
screen "0999_Service" 1280x800, template "Navigation"
   on GenerateScreen: SetTag("NavScreenChange", 5)
   on ClearScreen: SetTag("NavScreenChange", 0)
   Button "Button_3" at 326,104 size 451x32; TextOff 'Service'
   GraphicView "Graphic view_1" at 613,200 size 64x100; Picture "tank"
   GraphicView "Graphic view_2" at 385,180 size 144x140; Picture "Mcn"
   GraphicView "Graphic view_3" at 192,180 size 144x140; Picture "Machine"
   GraphicView "Graphic view_4" at 952,180 size 144x140; Picture "images_4"
   GraphicView "Graphic view_5" at 216,387 size 96x98; Picture "switch_off"
   GraphicView "Graphic view_6" at 781,224 size 116x60; Picture "Graphic_1"
   GraphicView "Graphic view_7" at 399,647 size 116x100; Picture "LARGESCALLEDVALUE"
   GraphicView "Graphic view_8" at 587,647 size 116x100; Picture "osiloskope_1"
   GraphicView "Graphic view_9" at 206,647 size 116x100; Picture "ethernet"
      Visibility <- "NavUserChange"
   Button "MixingHeadButton_1" at 565,182 size 160x136; TextOff 'Tank'; PictureOff "tank"
      on Click: ActivateScreen("0006_Tank", 0)
   Button "MixingHeadButton_3" at 944,182 size 160x136; TextOff 'Metering Pump'
      on Click: ActivateScreen("0004_Mixinghead", 0)
   Button "MixingHeadButton_2" at 184,182 size 160x136; TextOff 'General Machine'
      on Click: ActivateScreen("0021_Machine", 0)
   Button "MixingHeadButton_4" at 944,627 size 160x136; TextOff 'KM'; Authorization "User administration"
      Visibility <- "NavUserChange"
      on Click: ActivateScreen("2000_Configuration", 0)
   Button "MixingHeadButton_5" at 759,182 size 160x136; TextOff 'Mixinghead'
      on Click: ActivateScreen("0010_Pump", 0)
   Button "MixingHeadButton" at 377,182 size 160x136; TextOff 'Mixing Hydraulic'
      on Click: ActivateScreen("0002_MixingHeadHydraulic", 0)
   Button "MixingHeadButton_7" at 184,629 size 160x136; TextOff 'Network Setting'; Authorization "User administration"
      on Click: ActivateScreen("0014_Network Setting", 0)
      Visibility <- "NavUserChange"
   Button "MixingHeadButton_8" at 377,629 size 160x136; TextOff 'Large Scalled Values'
      on Click: ActivateScreen("0100_LargeScalledValues", 0); SetTag("NavScreenChange", 3); SetTag("LargeScalleValues Control", 1)
   Button "MixingHeadButton_9" at 565,629 size 160x136; TextOff 'Oscilloscope'
      on Click: ActivateScreen("0015_Oscilloscope", 0); SetTag("NavScreenChange", 2)
   Button "MixingHeadButton_10" at 184,368 size 160x136; TextOff 'Switch Menue'
      on Click: ActivateScreen("0009_Switch Menu", 0)
   Button "MixingHeadButton_11" at 759,623 size 160x136; TextOff 'Service & Solutions'
      on Click: ActivateScreen("9020_Service", 0)

screen "0016_Osciloscope Setting" 1280x800, template "Navigation"
   SymbolicIOField "Symbolic I/O field_11" at 704,218 size 160x30; TextOn '1'; TextOff '0'; TextList "oscilloscope_sensor_by_pump"
      Visibility <- "DB025_Oszilloskop_Graph{1}_Auswahl"
      ProcessValue <- "DB025_Oszilloskop_Graph{1}_Sensor"
   SymbolicIOField "Symbolic I/O field_15" at 704,270 size 160x30; TextOn '1'; TextOff '0'; TextList "oscilloscope_sensor_by_pump"
      Visibility <- "DB025_Oszilloskop_Graph{2}_Auswahl"
      ProcessValue <- "DB025_Oszilloskop_Graph{2}_Sensor"
   SymbolicIOField "Symbolic I/O field_19" at 704,322 size 160x30; TextOn '1'; TextOff '0'; TextList "oscilloscope_sensor_by_pump"
      ProcessValue <- "DB025_Oszilloskop_Graph{3}_Sensor"
      Visibility <- "DB025_Oszilloskop_Graph{3}_Auswahl"
   SymbolicIOField "Symbolic I/O field_23" at 704,374 size 160x30; TextOn '1'; TextOff '0'; TextList "oscilloscope_sensor_by_pump"
      ProcessValue <- "DB025_Oszilloskop_Graph{4}_Sensor"
      Visibility <- "DB025_Oszilloskop_Graph{4}_Auswahl"
   SymbolicIOField "Symbolic I/O field_27" at 704,426 size 160x30; TextOn '1'; TextOff '0'; TextList "oscilloscope_sensor_by_pump"
      ProcessValue <- "DB025_Oszilloskop_Graph{5}_Sensor"
      Visibility <- "DB025_Oszilloskop_Graph{5}_Auswahl"
   SymbolicIOField "Symbolic I/O field_31" at 704,478 size 160x30; TextOn '1'; TextOff '0'; TextList "oscilloscope_sensor_by_pump"
      ProcessValue <- "DB025_Oszilloskop_Graph{6}_Sensor"
      Visibility <- "DB025_Oszilloskop_Graph{6}_Auswahl"
   SymbolicIOField "Symbolic I/O field_35" at 704,530 size 160x30; TextOn '1'; TextOff '0'; TextList "oscilloscope_sensor_by_pump"
      ProcessValue <- "DB025_Oszilloskop_Graph{7}_Sensor"
      Visibility <- "DB025_Oszilloskop_Graph{7}_Auswahl"
   SymbolicIOField "Symbolic I/O field_39" at 704,582 size 160x30; TextOn '1'; TextOff '0'; TextList "oscilloscope_sensor_by_pump"
      ProcessValue <- "DB025_Oszilloskop_Graph{8}_Sensor"
      Visibility <- "DB025_Oszilloskop_Graph{8}_Auswahl"
   SymbolicIOField "Symbolic I/O field_12" at 704,218 size 160x30; TextOn '1'; TextOff '0'; TextList "oscilloscope_sensor_by_Tank"
      Visibility <- "DB025_Oszilloskop_Graph{1}_Auswahl"
      ProcessValue <- "DB025_Oszilloskop_Graph{1}_Sensor"
   SymbolicIOField "Symbolic I/O field_16" at 704,270 size 160x30; TextOn '1'; TextOff '0'; TextList "oscilloscope_sensor_by_Tank"
      Visibility <- "DB025_Oszilloskop_Graph{2}_Auswahl"
      ProcessValue <- "DB025_Oszilloskop_Graph{2}_Sensor"
   SymbolicIOField "Symbolic I/O field_20" at 704,322 size 160x30; TextOn '1'; TextOff '0'; TextList "oscilloscope_sensor_by_Tank"
      Visibility <- "DB025_Oszilloskop_Graph{3}_Auswahl"
      ProcessValue <- "DB025_Oszilloskop_Graph{3}_Sensor"
   SymbolicIOField "Symbolic I/O field_24" at 704,374 size 160x30; TextOn '1'; TextOff '0'; TextList "oscilloscope_sensor_by_Tank"
      Visibility <- "DB025_Oszilloskop_Graph{4}_Auswahl"
      ProcessValue <- "DB025_Oszilloskop_Graph{4}_Sensor"
   SymbolicIOField "Symbolic I/O field_28" at 704,426 size 160x30; TextOn '1'; TextOff '0'; TextList "oscilloscope_sensor_by_Tank"
      Visibility <- "DB025_Oszilloskop_Graph{5}_Auswahl"
      ProcessValue <- "DB025_Oszilloskop_Graph{5}_Sensor"
   SymbolicIOField "Symbolic I/O field_32" at 704,478 size 160x30; TextOn '1'; TextOff '0'; TextList "oscilloscope_sensor_by_Tank"
      Visibility <- "DB025_Oszilloskop_Graph{6}_Auswahl"
      ProcessValue <- "DB025_Oszilloskop_Graph{6}_Sensor"
   SymbolicIOField "Symbolic I/O field_36" at 704,530 size 160x30; TextOn '1'; TextOff '0'; TextList "oscilloscope_sensor_by_Tank"
      Visibility <- "DB025_Oszilloskop_Graph{7}_Auswahl"
      ProcessValue <- "DB025_Oszilloskop_Graph{7}_Sensor"
   SymbolicIOField "Symbolic I/O field_40" at 704,582 size 160x30; TextOn '1'; TextOff '0'; TextList "oscilloscope_sensor_by_Tank"
      Visibility <- "DB025_Oszilloskop_Graph{8}_Auswahl"
      ProcessValue <- "DB025_Oszilloskop_Graph{8}_Sensor"
   Button "Button_10" at 120,157 size 967x494; TextOff 'Text'
   Button "Button_3" at 326,104 size 451x32; TextOff 'Oscilloscope Settings'
   Button "Button_6" at 182,218 size 50x30; TextOff '1.'
   TextField "Text field_1" at 238,194 size 84x22; Text 'Selection'
   SymbolicIOField "Symbolic I/O field_1" at 238,218 size 160x30; TextOff '0'; TextOn '1'; TextList "oscilloscope_selection"
      ProcessValue <- "DB025_Oszilloskop_Graph{1}_Auswahl"
   Button "Button_1" at 182,270 size 50x30; TextOff '2.'
   TextField "Text field_2" at 238,246 size 84x22; Text 'Selection'
   SymbolicIOField "Symbolic I/O field_2" at 238,270 size 160x30; TextOn '1'; TextOff '0'; TextList "oscilloscope_selection"
      ProcessValue <- "DB025_Oszilloskop_Graph{2}_Auswahl"
   Button "Button_2" at 182,322 size 50x30; TextOff '3.'
   TextField "Text field_3" at 238,298 size 84x22; Text 'Selection'
   SymbolicIOField "Symbolic I/O field_3" at 238,322 size 160x30; TextOn '1'; TextOff '0'; TextList "oscilloscope_selection"
      ProcessValue <- "DB025_Oszilloskop_Graph{3}_Auswahl"
   Button "Button_4" at 182,374 size 50x30; TextOff '4.'
   TextField "Text field_4" at 238,350 size 84x22; Text 'Selection'
   SymbolicIOField "Symbolic I/O field_4" at 238,374 size 160x30; TextOn '1'; TextOff '0'; TextList "oscilloscope_selection"
      ProcessValue <- "DB025_Oszilloskop_Graph{4}_Auswahl"
   Button "Button_5" at 182,426 size 50x30; TextOff '5.'
   TextField "Text field_5" at 238,402 size 84x22; Text 'Selection'
   SymbolicIOField "Symbolic I/O field_5" at 238,426 size 160x30; TextOn '1'; TextOff '0'; TextList "oscilloscope_selection"
      ProcessValue <- "DB025_Oszilloskop_Graph{5}_Auswahl"
   Button "Button_7" at 182,478 size 50x30; TextOff '6.'
   TextField "Text field_6" at 238,454 size 84x22; Text 'Selection'
   SymbolicIOField "Symbolic I/O field_6" at 238,478 size 160x30; TextOn '1'; TextOff '0'; TextList "oscilloscope_selection"
      ProcessValue <- "DB025_Oszilloskop_Graph{6}_Auswahl"
   Button "Button_8" at 182,530 size 50x30; TextOff '7.'
   TextField "Text field_7" at 238,506 size 84x22; Text 'Selection'
   SymbolicIOField "Symbolic I/O field_7" at 238,530 size 160x30; TextOn '1'; TextOff '0'; TextList "oscilloscope_selection"
      ProcessValue <- "DB025_Oszilloskop_Graph{7}_Auswahl"
   Button "Button_9" at 182,582 size 50x30; TextOff '8.'
   TextField "Text field_8" at 238,558 size 84x22; Text 'Selection'
   SymbolicIOField "Symbolic I/O field_8" at 238,582 size 160x30; TextOn '1'; TextOff '0'; TextList "oscilloscope_selection"
      ProcessValue <- "DB025_Oszilloskop_Graph{8}_Auswahl"
   TextField "Text field_9" at 552,194 size 97x22; Text 'Component'
      Visibility <- "DB025_Oszilloskop_Graph{1}_Auswahl"
   TextField "Text field_10" at 744,194 size 68x22; Text 'Sensor'
      Visibility <- "DB025_Oszilloskop_Graph{1}_Auswahl"
   TextField "Text field_11" at 876,194 size 73x22; Text 'Scalling'
   TextField "Text field_12" at 968,194 size 80x22; Text 'DISPLAY'
   SymbolicIOField "Symbolic I/O field_9" at 528,218 size 160x30; TextOn '1'; TextOff '0'; TextList "oscilloscope_component_pump"
      ProcessValue <- "DB025_Oszilloskop_Graph{1}_Komponente"
      Visibility <- "DB025_Oszilloskop_Graph{1}_Auswahl"
   SymbolicIOField "Symbolic I/O field_10" at 704,218 size 160x30; TextOn '1'; TextOff '0'; TextList "oscilloscope_sensor_by_mh"
      ProcessValue <- "DB025_Oszilloskop_Graph{1}_Sensor"
      Visibility <- "DB025_Oszilloskop_Graph{1}_Auswahl"
   SymbolicIOField "Symbolic I/O field_13" at 528,270 size 160x30; TextOn '1'; TextOff '0'; TextList "oscilloscope_component_pump"
      ProcessValue <- "DB025_Oszilloskop_Graph{2}_Komponente"
      Visibility <- "DB025_Oszilloskop_Graph{2}_Auswahl"
   SymbolicIOField "Symbolic I/O field_14" at 704,270 size 160x30; TextOn '1'; TextOff '0'; TextList "oscilloscope_sensor_by_mh"
      Visibility <- "DB025_Oszilloskop_Graph{2}_Auswahl"
      ProcessValue <- "DB025_Oszilloskop_Graph{2}_Sensor"
   SymbolicIOField "Symbolic I/O field_17" at 528,322 size 160x30; TextOn '1'; TextOff '0'; TextList "oscilloscope_component_pump"
      ProcessValue <- "DB025_Oszilloskop_Graph{3}_Komponente"
      Visibility <- "DB025_Oszilloskop_Graph{3}_Auswahl"
   SymbolicIOField "Symbolic I/O field_18" at 704,322 size 160x30; TextOn '1'; TextOff '0'; TextList "oscilloscope_sensor_by_mh"
      ProcessValue <- "DB025_Oszilloskop_Graph{3}_Sensor"
      Visibility <- "DB025_Oszilloskop_Graph{3}_Auswahl"
   SymbolicIOField "Symbolic I/O field_21" at 528,374 size 160x30; TextOn '1'; TextOff '0'; TextList "oscilloscope_component_pump"
      ProcessValue <- "DB025_Oszilloskop_Graph{4}_Komponente"
      Visibility <- "DB025_Oszilloskop_Graph{4}_Auswahl"
   SymbolicIOField "Symbolic I/O field_22" at 704,374 size 160x30; TextOn '1'; TextOff '0'; TextList "oscilloscope_sensor_by_mh"
      ProcessValue <- "DB025_Oszilloskop_Graph{4}_Sensor"
      Visibility <- "DB025_Oszilloskop_Graph{4}_Auswahl"
   SymbolicIOField "Symbolic I/O field_25" at 528,426 size 160x30; TextOn '1'; TextOff '0'; TextList "oscilloscope_component_pump"
      ProcessValue <- "DB025_Oszilloskop_Graph{5}_Komponente"
      Visibility <- "DB025_Oszilloskop_Graph{5}_Auswahl"
   SymbolicIOField "Symbolic I/O field_26" at 704,426 size 160x30; TextOn '1'; TextOff '0'; TextList "oscilloscope_sensor_by_mh"
      Visibility <- "DB025_Oszilloskop_Graph{5}_Auswahl"
      ProcessValue <- "DB025_Oszilloskop_Graph{5}_Sensor"
   SymbolicIOField "Symbolic I/O field_29" at 528,478 size 160x30; TextOn '1'; TextOff '0'; TextList "oscilloscope_component_pump"
      ProcessValue <- "DB025_Oszilloskop_Graph{6}_Komponente"
      Visibility <- "DB025_Oszilloskop_Graph{6}_Auswahl"
   SymbolicIOField "Symbolic I/O field_30" at 704,478 size 160x30; TextOn '1'; TextOff '0'; TextList "oscilloscope_sensor_by_mh"
      ProcessValue <- "DB025_Oszilloskop_Graph{6}_Sensor"
      Visibility <- "DB025_Oszilloskop_Graph{6}_Auswahl"
   SymbolicIOField "Symbolic I/O field_33" at 528,530 size 160x30; TextOn '1'; TextOff '0'; TextList "oscilloscope_component_pump"
      ProcessValue <- "DB025_Oszilloskop_Graph{7}_Komponente"
      Visibility <- "DB025_Oszilloskop_Graph{7}_Auswahl"
   SymbolicIOField "Symbolic I/O field_34" at 704,530 size 160x30; TextOn '1'; TextOff '0'; TextList "oscilloscope_sensor_by_mh"
      ProcessValue <- "DB025_Oszilloskop_Graph{7}_Sensor"
      Visibility <- "DB025_Oszilloskop_Graph{7}_Auswahl"
   SymbolicIOField "Symbolic I/O field_37" at 528,582 size 160x30; TextOn '1'; TextOff '0'; TextList "oscilloscope_component_pump"
      ProcessValue <- "DB025_Oszilloskop_Graph{8}_Komponente"
      Visibility <- "DB025_Oszilloskop_Graph{8}_Auswahl"
   SymbolicIOField "Symbolic I/O field_38" at 704,582 size 160x30; TextOn '1'; TextOff '0'; TextList "oscilloscope_sensor_by_mh"
      ProcessValue <- "DB025_Oszilloskop_Graph{8}_Sensor"
      Visibility <- "DB025_Oszilloskop_Graph{8}_Auswahl"
   TextField "Text field_13" at 200,710 size 132x22; Text 'Starting Value / Starting Value:'
   TextField "Text field_14" at 200,752 size 93x22; Text 'End Value / End Value:'
   TextField "Text field_15" at 200,678 size 255x22; Text 'Scalling left,for selection 1-4'
   TextField "Text field_16" at 768,678 size 272x22; Text 'Scalling, right,for selection 5-8'
   TextField "Text field_17" at 768,710 size 132x22; Text 'Starting Value / Starting Value:'
   TextField "Text field_18" at 768,752 size 93x22; Text 'End Value / End Value:'
   TextField "Text field_19" at 876,246 size 73x22; Text 'Scalling'
   TextField "Text field_20" at 876,298 size 73x22; Text 'Scalling'
   TextField "Text field_21" at 876,350 size 73x22; Text 'Scalling'
   TextField "Text field_22" at 876,402 size 73x22; Text 'Scalling'
   TextField "Text field_23" at 876,454 size 73x22; Text 'Scalling'
   TextField "Text field_24" at 876,506 size 73x22; Text 'Scalling'
   TextField "Text field_25" at 876,558 size 73x22; Text 'Scalling'
   TextField "Text field_26" at 968,246 size 80x22; Text 'DISPLAY'
   TextField "Text field_27" at 968,298 size 80x22; Text 'DISPLAY'
   TextField "Text field_28" at 968,350 size 80x22; Text 'DISPLAY'
   TextField "Text field_29" at 968,402 size 80x22; Text 'DISPLAY'
   TextField "Text field_30" at 968,454 size 80x22; Text 'DISPLAY'
   TextField "Text field_31" at 968,506 size 80x22; Text 'DISPLAY'
   TextField "Text field_32" at 968,558 size 80x22; Text 'DISPLAY'
   TextField "Text field_33" at 552,246 size 97x22; Text 'Component'
      Visibility <- "DB025_Oszilloskop_Graph{2}_Auswahl"
   TextField "Text field_34" at 552,298 size 97x22; Text 'Component'
      Visibility <- "DB025_Oszilloskop_Graph{3}_Auswahl"
   TextField "Text field_35" at 552,350 size 97x22; Text 'Component'
      Visibility <- "DB025_Oszilloskop_Graph{4}_Auswahl"
   TextField "Text field_36" at 552,402 size 97x22; Text 'Component'
      Visibility <- "DB025_Oszilloskop_Graph{5}_Auswahl"
   TextField "Text field_37" at 552,454 size 97x22; Text 'Component'
      Visibility <- "DB025_Oszilloskop_Graph{6}_Auswahl"
   TextField "Text field_38" at 552,506 size 97x22; Text 'Component'
      Visibility <- "DB025_Oszilloskop_Graph{7}_Auswahl"
   TextField "Text field_39" at 552,558 size 97x22; Text 'Component'
      Visibility <- "DB025_Oszilloskop_Graph{8}_Auswahl"
   TextField "Text field_40" at 744,246 size 68x22; Text 'Sensor'
      Visibility <- "DB025_Oszilloskop_Graph{2}_Auswahl"
   TextField "Text field_41" at 744,298 size 68x22; Text 'Sensor'
      Visibility <- "DB025_Oszilloskop_Graph{3}_Auswahl"
   TextField "Text field_42" at 744,350 size 68x22; Text 'Sensor'
      Visibility <- "DB025_Oszilloskop_Graph{4}_Auswahl"
   TextField "Text field_43" at 744,402 size 68x22; Text 'Sensor'
      Visibility <- "DB025_Oszilloskop_Graph{5}_Auswahl"
   TextField "Text field_44" at 744,454 size 68x22; Text 'Sensor'
      Visibility <- "DB025_Oszilloskop_Graph{6}_Auswahl"
   TextField "Text field_45" at 744,506 size 68x22; Text 'Sensor'
      Visibility <- "DB025_Oszilloskop_Graph{7}_Auswahl"
   TextField "Text field_46" at 744,558 size 68x22; Text 'Sensor'
      Visibility <- "DB025_Oszilloskop_Graph{8}_Auswahl"
   IOField "I/O field_17" at 352,706 size 81x30; FormatPattern s9999
      ProcessValue <- "DB025_Oszilloskop_SkalierungGraphLinks_Startwert"
   IOField "I/O field_18" at 352,748 size 81x30; FormatPattern s9999
      ProcessValue <- "DB025_Oszilloskop_SkalierungGraphLinks_Ebdwert"
   IOField "I/O field_19" at 904,706 size 81x30; FormatPattern s9999
      ProcessValue <- "DB025_Oszilloskop_SkalierungGraphRechts_Startwert"
   IOField "I/O field_20" at 904,748 size 81x30; FormatPattern s9999
      ProcessValue <- "DB025_Oszilloskop_SkalierungGraphRechts_Ebdwert"
   IOField "Oscilloscope_Scalling_1" at 872,218 size 81x30; FormatPattern s999.9
      ProcessValue <- "DB025_Oszilloskop_Graph{1}_Skalierung"
   IOField "I/O field_3" at 872,270 size 81x30; FormatPattern s999.9
      ProcessValue <- "DB025_Oszilloskop_Graph{2}_Skalierung"
   IOField "I/O field_5" at 872,322 size 81x30; FormatPattern s999.9
      ProcessValue <- "DB025_Oszilloskop_Graph{3}_Skalierung"
   IOField "I/O field_7" at 872,374 size 81x30; FormatPattern s999.9
      ProcessValue <- "DB025_Oszilloskop_Graph{4}_Skalierung"
   IOField "I/O field_9" at 872,426 size 81x30; FormatPattern s999.9
      ProcessValue <- "DB025_Oszilloskop_Graph{5}_Skalierung"
   IOField "I/O field_11" at 872,478 size 81x30; FormatPattern s999.9
      ProcessValue <- "DB025_Oszilloskop_Graph{6}_Skalierung"
   IOField "I/O field_13" at 872,530 size 81x30; FormatPattern s999.9
      ProcessValue <- "DB025_Oszilloskop_Graph{7}_Skalierung"
   IOField "I/O field_15" at 872,582 size 81x30; FormatPattern s999.9
      ProcessValue <- "DB025_Oszilloskop_Graph{8}_Skalierung"
   IOField "I/O field_2" at 968,218 size 81x30; FormatPattern s999.9
      ProcessValue <- "DB025_Oszilloskop_Graph{1}_Wert"
   IOField "I/O field_4" at 968,270 size 81x30; FormatPattern s999.9
      ProcessValue <- "DB025_Oszilloskop_Graph{2}_Wert"
   IOField "I/O field_6" at 968,322 size 81x30; FormatPattern s999.9
      ProcessValue <- "DB025_Oszilloskop_Graph{3}_Wert"
   IOField "I/O field_8" at 968,374 size 81x30; FormatPattern s999.9
      ProcessValue <- "DB025_Oszilloskop_Graph{4}_Wert"
   IOField "I/O field_10" at 968,426 size 81x30; FormatPattern s999.9
      ProcessValue <- "DB025_Oszilloskop_Graph{5}_Wert"
   IOField "I/O field_12" at 968,478 size 81x30; FormatPattern s999.9
      ProcessValue <- "DB025_Oszilloskop_Graph{6}_Wert"
   IOField "I/O field_14" at 968,530 size 81x30; FormatPattern s999.9
      ProcessValue <- "DB025_Oszilloskop_Graph{7}_Wert"
   IOField "I/O field_16" at 968,582 size 81x30; FormatPattern s999.9
      ProcessValue <- "DB025_Oszilloskop_Graph{8}_Wert"
   SymbolicIOField "Symbolic I/O field_41" at 410,214 size 102x30; TextOn '1'; TextOff '0'; TextList "oscilloscope_MHnumber"
      Visibility <- "DB025_Oszilloskop_Graph{1}_Auswahl"
      ProcessValue <- "DB025_Oszilloskop_Graph{1}_Nummer"
   TextField "Text field_47" at 426,194 size 70x22; Text 'Number'
      Visibility <- "DB025_Oszilloskop_Graph{1}_Auswahl"
   SymbolicIOField "Symbolic I/O field_42" at 410,270 size 102x30; TextOn '1'; TextOff '0'; TextList "oscilloscope_MHnumber"
      Visibility <- "DB025_Oszilloskop_Graph{2}_Auswahl"
      ProcessValue <- "DB025_Oszilloskop_Graph{2}_Nummer"
   TextField "Text field_48" at 426,246 size 70x22; Text 'Number'
      Visibility <- "DB025_Oszilloskop_Graph{2}_Auswahl"
   SymbolicIOField "Symbolic I/O field_43" at 410,322 size 102x30; TextOn '1'; TextOff '0'; TextList "oscilloscope_MHnumber"
      Visibility <- "DB025_Oszilloskop_Graph{3}_Auswahl"
      ProcessValue <- "DB025_Oszilloskop_Graph{3}_Nummer"
   TextField "Text field_49" at 426,298 size 70x22; Text 'Number'
      Visibility <- "DB025_Oszilloskop_Graph{3}_Auswahl"
   SymbolicIOField "Symbolic I/O field_44" at 410,374 size 102x30; TextOn '1'; TextOff '0'; TextList "oscilloscope_MHnumber"
      Visibility <- "DB025_Oszilloskop_Graph{4}_Auswahl"
      ProcessValue <- "DB025_Oszilloskop_Graph{4}_Nummer"
   TextField "Text field_50" at 426,350 size 70x22; Text 'Number'
      Visibility <- "DB025_Oszilloskop_Graph{4}_Auswahl"
   SymbolicIOField "Symbolic I/O field_45" at 410,426 size 102x30; TextOn '1'; TextOff '0'; TextList "oscilloscope_MHnumber"
      Visibility <- "DB025_Oszilloskop_Graph{5}_Auswahl"
      ProcessValue <- "DB025_Oszilloskop_Graph{5}_Nummer"
   TextField "Text field_51" at 426,402 size 70x22; Text 'Number'
      Visibility <- "DB025_Oszilloskop_Graph{5}_Auswahl"
   SymbolicIOField "Symbolic I/O field_46" at 410,478 size 102x30; TextOn '1'; TextOff '0'; TextList "oscilloscope_MHnumber"
      Visibility <- "DB025_Oszilloskop_Graph{6}_Auswahl"
      ProcessValue <- "DB025_Oszilloskop_Graph{6}_Nummer"
   TextField "Text field_52" at 426,454 size 70x22; Text 'Number'
      Visibility <- "DB025_Oszilloskop_Graph{6}_Auswahl"
   SymbolicIOField "Symbolic I/O field_47" at 410,530 size 102x30; TextOn '1'; TextOff '0'; TextList "oscilloscope_MHnumber"
      Visibility <- "DB025_Oszilloskop_Graph{7}_Auswahl"
      ProcessValue <- "DB025_Oszilloskop_Graph{7}_Nummer"
   TextField "Text field_53" at 426,506 size 70x22; Text 'Number'
      Visibility <- "DB025_Oszilloskop_Graph{7}_Auswahl"
   SymbolicIOField "Symbolic I/O field_48" at 410,582 size 102x30; TextOn '1'; TextOff '0'; TextList "oscilloscope_MHnumber"
      Visibility <- "DB025_Oszilloskop_Graph{8}_Auswahl"
      ProcessValue <- "DB025_Oszilloskop_Graph{8}_Nummer"
   TextField "Text field_54" at 426,558 size 70x22; Text 'Number'
      Visibility <- "DB025_Oszilloskop_Graph{8}_Auswahl"
   SymbolicIOField "Symbolic I/O field_49" at 528,218 size 160x30; TextOn '1'; TextOff '0'; TextList "oscilloscope_component_tank"
      Visibility <- "DB025_Oszilloskop_Graph{1}_Auswahl"
      ProcessValue <- "DB025_Oszilloskop_Graph{1}_Komponente"
   SymbolicIOField "Symbolic I/O field_50" at 528,270 size 160x30; TextOn '1'; TextOff '0'; TextList "oscilloscope_component_tank"
      Visibility <- "DB025_Oszilloskop_Graph{2}_Auswahl"
      ProcessValue <- "DB025_Oszilloskop_Graph{2}_Komponente"
   SymbolicIOField "Symbolic I/O field_51" at 528,322 size 160x30; TextOn '1'; TextOff '0'; TextList "oscilloscope_component_tank"
      Visibility <- "DB025_Oszilloskop_Graph{3}_Auswahl"
      ProcessValue <- "DB025_Oszilloskop_Graph{3}_Komponente"
   SymbolicIOField "Symbolic I/O field_52" at 528,374 size 160x30; TextOn '1'; TextOff '0'; TextList "oscilloscope_component_tank"
      Visibility <- "DB025_Oszilloskop_Graph{4}_Auswahl"
      ProcessValue <- "DB025_Oszilloskop_Graph{4}_Komponente"
   SymbolicIOField "Symbolic I/O field_53" at 528,426 size 160x30; TextOn '1'; TextOff '0'; TextList "oscilloscope_component_tank"
      Visibility <- "DB025_Oszilloskop_Graph{5}_Auswahl"
      ProcessValue <- "DB025_Oszilloskop_Graph{5}_Komponente"
   SymbolicIOField "Symbolic I/O field_54" at 528,478 size 160x30; TextOn '1'; TextOff '0'; TextList "oscilloscope_component_tank"
      Visibility <- "DB025_Oszilloskop_Graph{6}_Auswahl"
      ProcessValue <- "DB025_Oszilloskop_Graph{6}_Komponente"
   SymbolicIOField "Symbolic I/O field_55" at 528,530 size 160x30; TextOn '1'; TextOff '0'; TextList "oscilloscope_component_tank"
      Visibility <- "DB025_Oszilloskop_Graph{7}_Auswahl"
      ProcessValue <- "DB025_Oszilloskop_Graph{7}_Komponente"
   SymbolicIOField "Symbolic I/O field_56" at 528,582 size 160x30; TextOn '1'; TextOff '0'; TextList "oscilloscope_component_tank"
      Visibility <- "DB025_Oszilloskop_Graph{8}_Auswahl"
      ProcessValue <- "DB025_Oszilloskop_Graph{8}_Komponente"

screen "0022_First_Screen" 1280x800, template "Navigation"
   on ClearScreen: "SettingShiftPlan"()
   TextField "KraussMaffei_Logo" at 328,360 size 712x120; Text 'Krauss Maffei'
   Button "b_First_Runtime" at 0,4 size 1272x790; TextOff 'Text'
      on Click: SetTag("First_Runtime_Rising_Control", 1); ActivateScreen("0017_Home Screen", 0); "FirstScreen_NavigationUpdate"()
      Visibility <- "First_Runtime_Rising_Control"

PopupScreen "Change DateTime" 620x248
   on GenerateScreen: "Move_Act_Time"()
   Button "Button_12" at 564,3 size 51x41; TextOff 'Text'; PictureOff "images (1)"
      on Press: function_efd93a16("Change DateTime", 0, 0, 0, -1, 1)
   TextField "Text field_1" at 191,7 size 258x29; Text 'Set Date & Time Clock / Set clock and date'
   Button "Button_3" at 135,186 size 338x41; TextOff 'SET'
      on Click: SetBit("TP-Bereichszeiger_Date_Time_Start_AG_Transfer")
   IOField "I/O field_1" at 43,73 size 56x32; FormatPattern 999
      ProcessValue <- "TP-Bereichszeiger_Date_Time_ActTime_DAY"
   IOField "I/O field_3" at 121,73 size 56x32; FormatPattern 999
      ProcessValue <- "TP-Bereichszeiger_Date_Time_ActTime_MONTH"
   IOField "I/O field_4" at 200,73 size 56x32; FormatPattern 99999
      ProcessValue <- "TP-Bereichszeiger_Date_Time_ActTime_YEAR"
   IOField "I/O field_6" at 351,73 size 56x32; FormatPattern 999
      ProcessValue <- "TP-Bereichszeiger_Date_Time_ActTime_HOUR"
   IOField "I/O field_7" at 429,73 size 56x32; FormatPattern 999
      ProcessValue <- "TP-Bereichszeiger_Date_Time_ActTime_MINUTE"
   IOField "I/O field_8" at 508,73 size 56x32; FormatPattern 999
      ProcessValue <- "TP-Bereichszeiger_Date_Time_ActTime_SECOND"
   IOField "I/O field_2" at 52,130 size 508x40; FormatPattern 99999999999999999999999999999999
      ProcessValue <- "TP-Bereichszeiger_Date_Time_SetTime"

screen "9021_Plc IO Monitor" 1280x800, template "Navigation"
   on GenerateScreen: SetTag("ServiceScreenControl", 9021)
   Button "Button_3" at 326,104 size 451x32; TextOff 'Plc Variabel / Service'
   IOField "Input_Byte" at 366,263 size 84x33; FormatPattern 99999
      ProcessValue <- "DB1025_Service_Set_Inputbyte"
   TextField "Text field_1" at 289,327 size 118x25; Text 'I .0'
   TextField "Text field_6" at 272,232 size 120x25; Text 'Input Byte :'
   IOField "Output_Byte" at 808,261 size 84x33; FormatPattern 99999
      ProcessValue <- "DB1025_Service_Set_Outputbyte"
   TextField "Text field_7" at 699,232 size 133x25; Text 'Output Byte :'
   Circle "Circle_1" at 409,324 size 32x32
      Appearance <- "DB1025_Service_State_Inputbyte"
   Circle "Circle_2" at 409,364 size 32x32
      Appearance <- "DB1025_Service_State_Inputbyte"
   Circle "Circle_3" at 409,404 size 32x32
      Appearance <- "DB1025_Service_State_Inputbyte"
   Circle "Circle_4" at 409,444 size 32x32
      Appearance <- "DB1025_Service_State_Inputbyte"
   Circle "Circle_5" at 409,484 size 32x32
      Appearance <- "DB1025_Service_State_Inputbyte"
   Circle "Circle_6" at 409,524 size 32x32
      Appearance <- "DB1025_Service_State_Inputbyte"
   Circle "Circle_7" at 409,564 size 32x32
      Appearance <- "DB1025_Service_State_Inputbyte"
   Circle "Circle_8" at 409,604 size 32x32
      Appearance <- "DB1025_Service_State_Inputbyte"
   TextField "Text field_11" at 749,327 size 121x25; Text 'Q .0'
   TextField "Text field_2" at 289,367 size 118x25; Text 'I .1'
   TextField "Text field_3" at 289,407 size 118x25; Text 'I .2'
   TextField "Text field_4" at 289,447 size 118x25; Text 'I .3'
   TextField "Text field_5" at 289,487 size 118x25; Text 'I .4'
   TextField "Text field_8" at 289,527 size 118x25; Text 'I .5'
   TextField "Text field_9" at 289,567 size 118x25; Text 'I .6'
   TextField "Text field_10" at 289,607 size 118x25; Text 'I .7'
   TextField "Text field_12" at 749,367 size 121x25; Text 'Q .1'
   TextField "Text field_13" at 749,407 size 121x25; Text 'Q .2'
   TextField "Text field_14" at 749,447 size 121x25; Text 'Q .3'
   TextField "Text field_15" at 749,487 size 121x25; Text 'Q .4'
   TextField "Text field_16" at 749,527 size 121x25; Text 'Q .5'
   TextField "Text field_17" at 749,567 size 121x25; Text 'Q .6'
   TextField "Text field_18" at 749,607 size 121x25; Text 'Q .7'
   Circle "Circle_17" at 861,324 size 32x32
      Appearance <- "DB1025_Service_State_Outputbyte"
   Circle "Circle_19" at 861,364 size 32x32
      Appearance <- "DB1025_Service_State_Outputbyte"
   Circle "Circle_20" at 861,404 size 32x32
      Appearance <- "DB1025_Service_State_Outputbyte"
   Circle "Circle_21" at 861,444 size 32x32
      Appearance <- "DB1025_Service_State_Outputbyte"
   Circle "Circle_22" at 861,484 size 32x32
      Appearance <- "DB1025_Service_State_Outputbyte"
   Circle "Circle_23" at 861,524 size 32x32
      Appearance <- "DB1025_Service_State_Outputbyte"
   Circle "Circle_24" at 861,564 size 32x32
      Appearance <- "DB1025_Service_State_Outputbyte"
   Circle "Circle_25" at 861,604 size 32x32
      Appearance <- "DB1025_Service_State_Outputbyte"
   Button "MixingHeadButton_6" at 219,696 size 60x60; TextOff 'PLC IO MONITOR'; PictureList "ico_plcio"
      on Click: ActivateScreen("9021_Plc IO Monitor", 0)
      Appearance <- "ServiceScreenControl"
      ProcessValue <- "ServiceScreenControl"
   Button "MixingHeadButton_2" at 308,696 size 60x60; TextOff 'PLC IO MONITOR Web'; PictureOff "ico"; PictureList "ico_Web"
      on Click: ActivateScreen("9022_Web Explorer", 0)
      ProcessValue <- "ServiceScreenControl"
      Appearance <- "ServiceScreenControl"
   Button "MixingHeadButton_3" at 397,696 size 60x60; TextOff 'PLC IO MONITOR smart'; PictureList "ico_Smart"
      on Click: ActivateScreen("9023_SmartClient", 0)
      Appearance <- "ServiceScreenControl"
      ProcessValue <- "ServiceScreenControl"
   Button "MixingHeadButton_5" at 397,696 size 60x60; TextOff 'PLC IO MONITOR smart'
      on Click: ActivateScreen("9023_SmartClient", 0)
      Appearance <- "ServiceScreenControl"
      ProcessValue <- "ServiceScreenControl"
   Button "MixingHeadButton_7" at 308,696 size 60x60; TextOff 'PLC IO MONITOR Web'
      on Click: ActivateScreen("9022_Web Explorer", 0)
      ProcessValue <- "ServiceScreenControl"
      Appearance <- "ServiceScreenControl"
   Button "MixingHeadButton_8" at 219,696 size 60x60; TextOff 'PLC IO MONITOR'
      on Click: ActivateScreen("9021_Plc IO Monitor", 0)
      Appearance <- "ServiceScreenControl"
      ProcessValue <- "ServiceScreenControl"
   Button "MixingHeadButton_9" at 1060,696 size 60x60; TextOff 'DIAGNOSTIC'; PictureOff "information"; PictureList "ico_information"
      on Click: ActivateScreen("9029_Information", 0)
      Appearance <- "ServiceScreenControl"
      ProcessValue <- "ServiceScreenControl"
   Button "MixingHeadButton_4" at 131,696 size 60x60; TextOff 'PLC IO MONITOR Service & Solutions'
      on Click: ActivateScreen("9020_Service", 0)
      Appearance <- "ServiceScreenControl"
   Button "MixingHeadButton_1" at 486,696 size 60x60; TextOff 'DIAGNOSTIC'; PictureOff "Graphic_29"
      on Click: ActivateScreen("9024_Diagnostic Overview", 0); function_ce3c6af1("9024_Diagnostic Overview", "System diagnostics view_1")
      Appearance <- "ServiceScreenControl"

screen "1000_General Machine Configuration" 1280x800, template "Navigation"
   TextField "Text field_1" at 227,206 size 203x25; Text 'Amount of machine :'
   TextField "Text field_2" at 227,240 size 230x25; Text 'Amount of component :'
   TextField "Text field_3" at 227,274 size 234x25; Text 'Amount of mixinghead :'
   TextField "Text field_4" at 227,308 size 166x25; Text 'Amount of tank :'
   TextField "Text field_5" at 227,342 size 251x25; Text 'Amount of mould carrier :'
   TextField "Text field_6" at 227,376 size 194x25; Text 'Amount of module :'
   TextField "Text field_7" at 227,440 size 193x25; Text 'Amount of Station :'
   TextField "Text field_8" at 227,594 size 318x25; Text 'Program number from interface :'
   TextField "Text field_9" at 227,631 size 347x25; Text 'Mixinghead number from interface :'
   IOField "I/O field_2" at 519,203 size 166x30; Authorization "User administration"; FormatPattern 9999
      ProcessValue <- "DB790_PlantParameter_AmountMachine"
   IOField "Amount_Of_Component" at 519,237 size 166x30; Authorization "User administration"; FormatPattern 9999
      ProcessValue <- "DB790_PlantParameter_AmountMeteringUnits"
   IOField "I/O field_3" at 519,271 size 166x30; Authorization "User administration"; FormatPattern 9999
      ProcessValue <- "DB790_PlantParameter_AmountMH"
   IOField "I/O field_4" at 519,305 size 166x30; Authorization "User administration"; FormatPattern 9999
      ProcessValue <- "DB790_PlantParameter_AmountTank"
   IOField "I/O field_5" at 519,339 size 166x30; Authorization "User administration"; FormatPattern 9999
      ProcessValue <- "DB790_PlantParameter_AmountMouldCarrier"
   IOField "I/O field_6" at 519,373 size 166x30; Authorization "User administration"; FormatPattern 9999
      ProcessValue <- "DB790_PlantParameter_AmountProCanModul"
   IOField "I/O field_7" at 519,437 size 166x30; Authorization "User administration"; FormatPattern 9999
      ProcessValue <- "DB790_PlantParameter_AmountToolStation"
   Button "Check_Mhydraulic_Prog_number_interface" at 640,591 size 45x30; TextOff 'Text'; PictureOff "download"; PictureList "Check_Uncheck"; Authorization "User administration"
      ProcessValue <- "DB790_PlantParameter_Bit_ProgrammNofromInterface"
      on Click: InvertBit("DB790_PlantParameter_Bit_ProgrammNofromInterface")
   Button "Check_Mhydraulic_MH_number_interface" at 640,628 size 45x30; TextOff 'Text'; PictureOff "download"; PictureList "Check_Uncheck"; Authorization "User administration"
      ProcessValue <- "DB790_PlantParameter_Bit_MHNofromInterface"
      on Click: InvertBit("DB790_PlantParameter_Bit_MHNofromInterface")
   TextField "Text field_10" at 462,118 size 357x29; Text 'General Machine Configuration'
   TextField "Text field_11" at 227,536 size 193x25; Text 'Amount of Station : / Amount of Robots :'
      Visibility <- "DB704_MH_Value_Mixinghead{0}_Conf_IntWithRobot"
   IOField "I/O field_1" at 519,533 size 166x30; Authorization "User administration"; FormatPattern 9999
      ProcessValue <- "DB790_PlantParameter_AmountRobots"
      Visibility <- "DB704_MH_Value_Mixinghead{0}_Conf_IntWithRobot"

screen "2000_Configuration" 1280x800, template "Navigation"
   Button "Button_3" at 326,104 size 451x32; TextOff 'Configuration'
   Button "Button_1" at 150,238 size 251x40; TextOff 'ProNet Mixinghead / ProNet MH digital'
      on Press: ActivateScreen("2004_ProNet MH digital", 0)
   Button "Button_2" at 150,293 size 251x40; TextOff 'Pronet Cleaning Piston / ProNet CP digital'
      on Press: ActivateScreen("2003_ProNet CP digital", 0)
   Button "Button_4" at 150,348 size 251x40; TextOff 'Pronet Analog Input 1 / ProNet analog input'
      on Press: ActivateScreen("2001_ProNet analog input", 0)
   Button "Button_5" at 150,403 size 251x40; TextOff 'Pronet Analog Input 2 / ProNet temperature input'
      on Press: ActivateScreen("2005_ProNet temperature input", 0)
   Button "Button_6" at 150,458 size 251x40; TextOff 'Pronet Flow control / ProNet flow control'
      on Press: ActivateScreen("2002_ProNet Flow control", 0)
   Button "Button_7" at 150,513 size 251x40; TextOff 'Pronet Nozzle Control 1 / ProNet nozzle configuration'
      on Press: ActivateScreen("2006_ProNet Nozzle configuration", 0)
   Button "Button_8" at 150,568 size 251x40; TextOff 'Pronet Nozzle Control 2 / ProNet nozzle times'
      on Press: ActivateScreen("2007_ProNet Nozzle times", 0)
   Button "Button_9" at 150,623 size 251x40; TextOff 'ProNet Diagnose IO'
      on Click: ActivateScreen("2009_ProNet Diagnose IO", 0)
   Button "Button_10" at 421,243 size 296x40; TextOff 'Config PV Tank'
      on Press: ActivateScreen("1001_Process Value Tank", 0)
   Button "Button_11" at 421,293 size 296x40; TextOff 'Config PV Metering'
      on Press: ActivateScreen("1003_Process Value MeteringUnit", 0)
   Button "Button_12" at 421,343 size 296x40; TextOff 'Config PV MixingHead'
      on Press: ActivateScreen("1002_Process Value Mixing Head", 0)
   Button "Button_13" at 421,393 size 296x40; TextOff 'Config PV MH Inerting'
      on Press: ActivateScreen("1005_Process Value MH Inerting", 0)
   Button "Button_14" at 150,158 size 203x40; TextOff 'ProNet Module Config'
   Button "Button_15" at 421,158 size 203x40; TextOff 'Procces Values'

screen "1001_Process Value Tank" 1280x800, template "Navigation"
   on GenerateScreen: SetBit("DB702_Tank_Value_Read")
   TextField "Text field_12" at 526,557 size 53x25; Text '[ C ]'
   TextField "Text field_13" at 534,556 size 36x18; Text 'O'
   Group "Group_1" at 118,177 size 1041x522
   TextField "Text field_1" at 319,143 size 232x29; Text 'Process values tank'
   TextField "Text field_2" at 243,258 size 112x25; Text 'Module No.'
   TextField "Text field_3" at 243,306 size 81x25; Text 'Address'
   TextField "Text field_4" at 243,354 size 64x25; Text 'Offset'
   TextField "Text field_5" at 243,402 size 96x25; Text 'Multiplier'
   TextField "Text field_6" at 243,450 size 174x25; Text 'Min. Value Sensor'
   TextField "Text field_7" at 243,498 size 178x25; Text 'Max. Value Sensor'
   TextField "Text field_8" at 243,606 size 123x25; Text 'Actual Value'
   TextField "Text field_9" at 490,208 size 125x25; Text 'Temperature'
   TextField "Text field_10" at 709,208 size 55x25; Text 'Level'
   TextField "Text field_11" at 867,208 size 107x25; Text 'Nucleation'
   IOField "ModuleNo_Temperature_PV_Tank" at 481,255 size 142x30; Authorization "User administration"; FormatPattern 99999
      ProcessValue <- "DB602_PV_Tank_Tank{0}_Temp_PV_Conf_ActV_ModulNo"
   IOField "I/O field_2" at 481,303 size 142x30; Authorization "User administration"; FormatPattern 99999
      ProcessValue <- "DB602_PV_Tank_Tank{0}_Temp_PV_Conf_ActV_Address"
   IOField "I/O field_3" at 481,351 size 142x30; Authorization "User administration"; FormatPattern 99999
      ProcessValue <- "DB602_PV_Tank_Tank{0}_Temp_PV_Conf_ActV_OffsetSignal"
   IOField "I/O field_4" at 481,399 size 142x30; Authorization "User administration"; FormatPattern 9999.999
      ProcessValue <- "DB602_PV_Tank_Tank{0}_Temp_PV_Conf_ActV_Multiplier"
   IOField "I/O field_5" at 481,447 size 142x30; Authorization "User administration"; FormatPattern 9999999
      ProcessValue <- "DB602_PV_Tank_Tank{0}_Temp_PV_Conf_ActV_MinValueSensor"
   IOField "I/O field_6" at 481,495 size 142x30; Authorization "User administration"; FormatPattern 9999999
      ProcessValue <- "DB602_PV_Tank_Tank{0}_Temp_PV_Conf_ActV_MaxValueSensor"
   IOField "I/O field_7" at 514,603 size 77x30; FormatPattern 999.9
      ProcessValue <- "DB602_PV_Tank_Tank{0}_Temp_PV_ActV_Value"
   Group "Group" at 526,556 size 53x26
   TextField "Text field_14" at 714,557 size 46x25; Text '[%]'
   TextField "Text field_15" at 898,557 size 46x25; Text '[%]'
   IOField "I/O field_8" at 665,254 size 142x30; Authorization "User administration"; FormatPattern 99999
      ProcessValue <- "DB602_PV_Tank_Tank{0}_Level_PV_Conf_ActV_ModulNo"
   IOField "I/O field_9" at 665,302 size 142x30; Authorization "User administration"; FormatPattern 99999
      ProcessValue <- "DB602_PV_Tank_Tank{0}_Level_PV_Conf_ActV_Address"
   IOField "I/O field_10" at 665,350 size 142x30; Authorization "User administration"; FormatPattern 99999
      ProcessValue <- "DB602_PV_Tank_Tank{0}_Level_PV_Conf_ActV_OffsetSignal"
   IOField "I/O field_11" at 665,398 size 142x30; Authorization "User administration"; FormatPattern 9999.999
      ProcessValue <- "DB602_PV_Tank_Tank{0}_Level_PV_Conf_ActV_Multiplier"
   IOField "I/O field_12" at 665,446 size 142x30; Authorization "User administration"; FormatPattern 9999999
      ProcessValue <- "DB602_PV_Tank_Tank{0}_Level_PV_Conf_ActV_MinValueSensor"
   IOField "I/O field_13" at 665,494 size 142x30; Authorization "User administration"; FormatPattern 9999999
      ProcessValue <- "DB602_PV_Tank_Tank{0}_Level_PV_Conf_ActV_MaxValueSensor"
   IOField "I/O field_14" at 849,253 size 142x30; Authorization "User administration"; FormatPattern 99999
      ProcessValue <- "DB602_PV_Tank_Tank{0}_Nucleation_PV_Conf_ActV_ModulNo"
   IOField "I/O field_15" at 849,301 size 142x30; Authorization "User administration"; FormatPattern 99999
      ProcessValue <- "DB602_PV_Tank_Tank{0}_Nucleation_PV_Conf_ActV_Address"
   IOField "I/O field_16" at 849,349 size 142x30; Authorization "User administration"; FormatPattern 99999
      ProcessValue <- "DB602_PV_Tank_Tank{0}_Nucleation_PV_Conf_ActV_OffsetSignal"
   IOField "I/O field_17" at 849,397 size 142x30; Authorization "User administration"; FormatPattern 9999.999
      ProcessValue <- "DB602_PV_Tank_Tank{0}_Nucleation_PV_Conf_ActV_Multiplier"
   IOField "I/O field_18" at 849,445 size 142x30; Authorization "User administration"; FormatPattern 9999999
      ProcessValue <- "DB602_PV_Tank_Tank{0}_Nucleation_PV_Conf_ActV_MinValueSensor"
   IOField "I/O field_19" at 849,493 size 142x30; Authorization "User administration"; FormatPattern 9999999
      ProcessValue <- "DB602_PV_Tank_Tank{0}_Nucleation_PV_Conf_ActV_MaxValueSensor"
   IOField "I/O field_20" at 698,602 size 77x30; FormatPattern 999.9
      ProcessValue <- "DB602_PV_Tank_Tank{0}_Level_PV_ActV_Value"
   IOField "I/O field_21" at 882,601 size 77x30; FormatPattern 999.9
      ProcessValue <- "DB602_PV_Tank_Tank{0}_Nucleation_PV_ActV_Value"
   SymbolicIOField "Symbolic I/O field_1" at 326,104 size 451x32; TextOff '0'; TextOn '1'; TextList "Tank_IOField"
      ProcessValue <- "DB612_Tank_State.ReadDeviceNo"
   Button "b_Incress_PV_Tank" at 786,104 size 46x32; TextOff 'Text'; PictureOff "NEXT"
      on Click: function_dd21b452("DB612_Tank_State.ReadDeviceNo", 1)
   Button "b_Decress_PV_Tank" at 271,104 size 46x32; TextOff 'Text'; PictureOff "BEFORE"
      on Click: function_b9b71300("DB612_Tank_State.ReadDeviceNo", 1)
      ObjectEnable <- "DB612_Tank_State.ReadDeviceNo"

screen "1003_Process Value MeteringUnit" 1280x800, template "Navigation"
   on GenerateScreen: SetBit("DB613_Komponent_State_Write"); SetBit("DB608_PV_Metering_Read")
   TextField "Text field_12" at 421,523 size 53x25; Text '[ C ]'
   TextField "Text field_13" at 429,522 size 36x18; Text 'O'
   TextField "Text field_20" at 1052,529 size 53x25; Text '[ C ]'
   TextField "Text field_21" at 1060,528 size 36x18; Text 'O'
   Group "Group_2" at 100,184 size 1076x496
   TextField "Text field_1" at 484,147 size 309x27; Text 'Process values metering unit'
   TextField "Text field_2" at 138,242 size 112x25; Text 'Module No.'
   TextField "Text field_3" at 138,290 size 81x25; Text 'Address'
   TextField "Text field_4" at 138,338 size 64x25; Text 'Offset'
   TextField "Text field_5" at 138,386 size 96x25; Text 'Multiplier'
   TextField "Text field_6" at 138,434 size 174x25; Text 'Min. Value Sensor'
   TextField "Text field_7" at 138,482 size 178x25; Text 'Max. Value Sensor'
   TextField "Text field_8" at 138,564 size 123x25; Text 'Actual Value'
   TextField "Text field_9" at 382,206 size 125x25; Text 'Temperature'
   TextField "Text field_10" at 531,206 size 124x25; Text 'Pre Pressure'
   TextField "Text field_11" at 718,206 size 87x25; Text 'Pressure'
   IOField "Pronet_PV_MU_ModulNo_Temperature" at 373,240 size 142x30; Authorization "User administration"; FormatPattern 9999999
      ProcessValue <- "DB608_PV_Metering_Metering{0}_Temperature_PV_Conf_ActV_ModulNo"
   IOField "I/O field_2" at 373,288 size 142x30; Authorization "User administration"; FormatPattern 9999999
      ProcessValue <- "DB608_PV_Metering_Metering{0}_Temperature_PV_Conf_ActV_Address"
   IOField "I/O field_3" at 373,336 size 142x30; Authorization "User administration"; FormatPattern 9999999
      ProcessValue <- "DB608_PV_Metering_Metering{0}_Temperature_PV_Conf_ActV_OffsetSignal"
   IOField "I/O field_4" at 373,384 size 142x30; Authorization "User administration"; FormatPattern s99999.999
      ProcessValue <- "DB608_PV_Metering_Metering{0}_Temperature_PV_Conf_ActV_Multiplier"
   IOField "I/O field_5" at 373,432 size 142x30; Authorization "User administration"; FormatPattern s9999999
      ProcessValue <- "DB608_PV_Metering_Metering{0}_Temperature_PV_Conf_ActV_MinValueSensor"
   IOField "I/O field_6" at 373,480 size 142x30; Authorization "User administration"; FormatPattern s9999999
      ProcessValue <- "DB608_PV_Metering_Metering{0}_Temperature_PV_Conf_ActV_MaxValueSensor"
   IOField "I/O field_7" at 373,562 size 142x30; Authorization "User administration"; FormatPattern 99999.9
      ProcessValue <- "DB608_PV_Metering_Metering{0}_Temperature_PV_ActV_Value"
   Group "Group" at 421,522 size 53x26
   TextField "Text field_14" at 579,523 size 54x25; Text '[bar]'
   TextField "Text field_15" at 733,526 size 54x25; Text '[bar]'
   IOField "I/O field_8" at 531,240 size 142x30; Authorization "User administration"; FormatPattern 9999999
      ProcessValue <- "DB608_PV_Metering_Metering{0}_Pre_Pressure_PV_Conf_ActV_ModulNo"
   IOField "I/O field_9" at 531,288 size 142x30; Authorization "User administration"; FormatPattern 9999999
      ProcessValue <- "DB608_PV_Metering_Metering{0}_Pre_Pressure_PV_Conf_ActV_Address"
   IOField "I/O field_10" at 531,336 size 142x30; Authorization "User administration"; FormatPattern 9999999
      ProcessValue <- "DB608_PV_Metering_Metering{0}_Pre_Pressure_PV_Conf_ActV_OffsetSignal"
   IOField "I/O field_11" at 531,384 size 142x30; Authorization "User administration"; FormatPattern s99999.999
      ProcessValue <- "DB608_PV_Metering_Metering{0}_Pre_Pressure_PV_Conf_ActV_Multiplier"
   IOField "I/O field_12" at 531,432 size 142x30; Authorization "User administration"; FormatPattern s9999999
      ProcessValue <- "DB608_PV_Metering_Metering{0}_Pre_Pressure_PV_Conf_ActV_MinValueSensor"
   IOField "I/O field_13" at 531,480 size 142x30; Authorization "User administration"; FormatPattern s9999999
      ProcessValue <- "DB608_PV_Metering_Metering{0}_Pre_Pressure_PV_Conf_ActV_MaxValueSensor"
   IOField "I/O field_14" at 690,240 size 142x30; Authorization "User administration"; FormatPattern 9999999
      ProcessValue <- "DB608_PV_Metering_Metering{0}_Pressure_PV_Conf_ActV_ModulNo"
   IOField "I/O field_15" at 690,288 size 142x30; Authorization "User administration"; FormatPattern 9999999
      ProcessValue <- "DB608_PV_Metering_Metering{0}_Pressure_PV_Conf_ActV_Address"
   IOField "I/O field_16" at 690,336 size 142x30; Authorization "User administration"; FormatPattern 9999999
      ProcessValue <- "DB608_PV_Metering_Metering{0}_Pressure_PV_Conf_ActV_OffsetSignal"
   IOField "I/O field_17" at 690,384 size 142x30; Authorization "User administration"; FormatPattern s99999.999
      ProcessValue <- "DB608_PV_Metering_Metering{0}_Pressure_PV_Conf_ActV_Multiplier"
   IOField "I/O field_18" at 690,432 size 142x30; Authorization "User administration"; FormatPattern s9999999
      ProcessValue <- "DB608_PV_Metering_Metering{0}_Pressure_PV_Conf_ActV_MinValueSensor"
   IOField "I/O field_19" at 690,480 size 142x30; Authorization "User administration"; FormatPattern s9999999
      ProcessValue <- "DB608_PV_Metering_Metering{0}_Pressure_PV_Conf_ActV_MaxValueSensor"
   IOField "I/O field_20" at 531,562 size 142x30; Authorization "User administration"; FormatPattern 99999.9
      ProcessValue <- "DB608_PV_Metering_Metering{0}_Pre_Pressure_PV_ActV_Value"
   IOField "I/O field_21" at 690,562 size 142x30; Authorization "User administration"; FormatPattern 99999.9
      ProcessValue <- "DB608_PV_Metering_Metering{0}_Pressure_PV_ActV_Value"
   SymbolicIOField "Symbolic I/O field_1" at 326,104 size 451x32; TextOn '1'; TextOff '0'; TextList "Tank_IOField"
      ProcessValue <- "DB613_Komponent_State_ReadDeviceNo"
   TextField "Text field_16" at 894,206 size 50x25; Text 'Flow'
   TextField "Text field_17" at 1019,206 size 125x25; Text 'HP HeatExch'
   IOField "I/O field_22" at 848,288 size 142x30; Authorization "User administration"; FormatPattern 9999999
      ProcessValue <- "DB608_PV_Metering_Metering{0}_Flow_PV_Conf_ActV_Address"
   IOField "I/O field_23" at 1010,240 size 142x30; Authorization "User administration"; FormatPattern 9999999
      ProcessValue <- "DB608_PV_Metering_HeatexchangerHP{0}_PV_Conf_ActV_ModulNo"
   IOField "I/O field_24" at 1010,288 size 142x30; Authorization "User administration"; FormatPattern 9999999
      ProcessValue <- "DB608_PV_Metering_HeatexchangerHP{0}_PV_Conf_ActV_Address"
   IOField "I/O field_25" at 1010,336 size 142x30; Authorization "User administration"; FormatPattern 9999999
      ProcessValue <- "DB608_PV_Metering_HeatexchangerHP{0}_PV_Conf_ActV_OffsetSignal"
   IOField "I/O field_26" at 1010,384 size 142x30; Authorization "User administration"; FormatPattern s99999.999
      ProcessValue <- "DB608_PV_Metering_HeatexchangerHP{0}_PV_Conf_ActV_Multiplier"
   IOField "I/O field_27" at 1010,432 size 142x30; Authorization "User administration"; FormatPattern s9999999
      ProcessValue <- "DB608_PV_Metering_HeatexchangerHP{0}_PV_Conf_ActV_MinValueSensor"
   IOField "I/O field_28" at 1010,480 size 142x30; Authorization "User administration"; FormatPattern s9999999
      ProcessValue <- "DB608_PV_Metering_HeatexchangerHP{0}_PV_Conf_ActV_MaxValueSensor"
   IOField "I/O field_29" at 1010,562 size 142x30; Authorization "User administration"; FormatPattern 99999.9
      ProcessValue <- "DB608_PV_Metering_HeatexchangerHP{0}_PV_ActV_Value"
   TextField "Text field_19" at 894,528 size 56x25; Text '[g/s]'
   IOField "I/O field_30" at 848,562 size 142x30; Authorization "User administration"; FormatPattern 99999.99
      ProcessValue <- "DB608_PV_Metering_Metering{0}_Flow_PV_ActV_Value"
   Group "Group_1" at 1052,528 size 53x26
   IOField "I/O field_31" at 373,603 size 142x30; Authorization "User administration"; FormatPattern s9999999
      ProcessValue <- "DB608_PV_Metering_Metering{0}_Temperature_PV_Conf_ActV_MaxSignalResolution"
   IOField "I/O field_32" at 531,602 size 142x30; Authorization "User administration"; FormatPattern s9999999
      ProcessValue <- "DB608_PV_Metering_Metering{0}_Pre_Pressure_PV_Conf_ActV_MaxSignalResolution"
   IOField "I/O field_33" at 690,601 size 142x30; Authorization "User administration"; FormatPattern s9999999
      ProcessValue <- "DB608_PV_Metering_Metering{0}_Pressure_PV_Conf_ActV_MaxSignalResolution"
   IOField "I/O field_34" at 1010,604 size 142x30; Authorization "User administration"; FormatPattern s9999999
      ProcessValue <- "DB608_PV_Metering_HeatexchangerHP{0}_PV_Conf_ActV_MaxSignalResolution"
   TextField "Text field_18" at 138,606 size 216x25; Text 'Max Signal Resolution'
   TextField "Text field_22" at 138,691 size 81x25; Text 'Address'
   TextField "Text field_23" at 138,723 size 64x25; Text 'Offset'
   TextField "Text field_24" at 138,758 size 96x25; Text 'Multiplier'
   TextField "Text field_25" at 382,691 size 371x25; Text 'Address Number PLC or ProCan Chanel'
   TextField "Text field_26" at 382,723 size 321x25; Text 'Value to add the calculated value'
   TextField "Text field_27" at 382,748 size 364x25; Text 'conversion value for the actual value'
   TextField "Text field_28" at 382,770 size 300x25; Text '(signal detail/max.value x100)'
   Button "b_Incress_PV_MU" at 786,104 size 46x32; TextOff 'Text'; PictureOff "NEXT"
      on Click: function_dd21b452("DB613_Komponent_State_ReadDeviceNo", 1)
   Button "b_Decress_PV_MU" at 272,104 size 46x32; TextOff 'Text'; PictureOff "BEFORE"
      on Click: function_b9b71300("DB613_Komponent_State_ReadDeviceNo", 1)

